   266: 'Carrier 04 Safe Output Card Fault', class No Acknowledgement, trigger "DB302_HMI_Faults_Carrier4_Faults_0" bit 9
   267: 'Carrier 04 Standard Input Card Fault', class No Acknowledgement, trigger "DB302_HMI_Faults_Carrier4_Faults_0" bit 10
   268: 'Carrier 04 Standard Output Card Fault', class No Acknowledgement, trigger "DB302_HMI_Faults_Carrier4_Faults_0" bit 11
   269: 'Carrier 04 Encoder Position Fault', class No Acknowledgement, trigger "DB302_HMI_Faults_Carrier4_Faults_0" bit 12
   270: 'Carrier 04 Encoder Internal Error', class No Acknowledgement, trigger "DB302_HMI_Faults_Carrier4_Faults_0" bit 13
   271: 'Carrier 04 Encoder Comm Fault', class No Acknowledgement, trigger "DB302_HMI_Faults_Carrier4_Faults_0" bit 14
   272: 'Carrier 04 HMI Comm Fault', class No Acknowledgement, trigger "DB302_HMI_Faults_Carrier4_Faults_0" bit 15
   273: 'Carrier 04 Crash Detection Fault', class No Acknowledgement, trigger "DB302_HMI_Faults_Carrier4_Faults_1" bit 0
   274: 'Carrier 04 Carrier Number Invalid', class No Acknowledgement, trigger "DB302_HMI_Faults_Carrier4_Faults_1" bit 1
   275: 'Carrier 04 Drive: PROFINET configuration error', class No Acknowledgement, trigger "DB302_HMI_Faults_Carrier4_Faults_1" bit 2
   276: 'Carrier 04 Drive: Error internal communications', class No Acknowledgement, trigger "DB302_HMI_Faults_Carrier4_Faults_1" bit 3
   277: 'Carrier 04 Drive: Motor overtemperature', class No Acknowledgement, trigger "DB302_HMI_Faults_Carrier4_Faults_1" bit 4
   278: 'Carrier 04 Drive: Motor overcurrent', class No Acknowledgement, trigger "DB302_HMI_Faults_Carrier4_Faults_1" bit 5
   279: 'Carrier 04 Drive: Infeed or power unit not ready', class No Acknowledgement, trigger "DB302_HMI_Faults_Carrier4_Faults_1" bit 6
   280: 'Carrier 04 Drive: Short-circuit/ground fault detected', class No Acknowledgement, trigger "DB302_HMI_Faults_Carrier4_Faults_1" bit 7
   281: 'Carrier 04 Drive: PROFINET Setpoint timeout', class No Acknowledgement, trigger "DB302_HMI_Faults_Carrier4_Faults_1" bit 8
   282: 'Carrier 04 Power unit: Overcurrent', class No Acknowledgement, trigger "DB302_HMI_Faults_Carrier4_Faults_1" bit 9
   283: 'Carrier 04 Power unit: DC link voltage overvoltage', class No Acknowledgement, trigger "DB302_HMI_Faults_Carrier4_Faults_1" bit 10
   284: 'Carrier 04 Power unit: DC link voltage undervoltage', class No Acknowledgement, trigger "DB302_HMI_Faults_Carrier4_Faults_1" bit 11
   285: 'Carrier 04 Power unit: Line phase failure in main circuit', class No Acknowledgement, trigger "DB302_HMI_Faults_Carrier4_Faults_1" bit 12
   286: 'Carrier 04 Power unit: Phase failure motor cable', class No Acknowledgement, trigger "DB302_HMI_Faults_Carrier4_Faults_1" bit 13
   287: 'Carrier 04 Power unit: Ground fault', class No Acknowledgement, trigger "DB302_HMI_Faults_Carrier4_Faults_1" bit 14
   288: 'Spare_Fault_288', class No Acknowledgement, trigger "DB302_HMI_Faults_Carrier4_Faults_1" bit 15
   289: 'Carrier 04 Motion Off Fault', class No Acknowledgement, trigger "DB302_HMI_Faults_Carrier4_Faults_2" bit 0
   290: 'Carrier 04 Motion On Fault', class No Acknowledgement, trigger "DB302_HMI_Faults_Carrier4_Faults_2" bit 1
   291: 'Carrier 04 Spacing Fault', class No Acknowledgement, trigger "DB302_HMI_Faults_Carrier4_Faults_2" bit 2
   292: 'Carrier 04 Duplicate Carrier Number Fault', class No Acknowledgement, trigger "DB302_HMI_Faults_Carrier4_Faults_2" bit 3
   293: 'Spare_Fault_293', class No Acknowledgement, trigger "DB302_HMI_Faults_Carrier4_Faults_2" bit 4
   294: 'Spare_Fault_294', class No Acknowledgement, trigger "DB302_HMI_Faults_Carrier4_Faults_2" bit 5
   295: 'Spare_Fault_295', class No Acknowledgement, trigger "DB302_HMI_Faults_Carrier4_Faults_2" bit 6
   296: 'Spare_Fault_296', class No Acknowledgement, trigger "DB302_HMI_Faults_Carrier4_Faults_2" bit 7
   297: 'Spare_Fault_297', class No Acknowledgement, trigger "DB302_HMI_Faults_Carrier4_Faults_2" bit 8
   298: 'Spare_Fault_298', class No Acknowledgement, trigger "DB302_HMI_Faults_Carrier4_Faults_2" bit 9
   299: 'Spare_Fault_299', class No Acknowledgement, trigger "DB302_HMI_Faults_Carrier4_Faults_2" bit 10
   300: 'Spare_Fault_300', class No Acknowledgement, trigger "DB302_HMI_Faults_Carrier4_Faults_2" bit 11
   301: 'Spare_Fault_301', class No Acknowledgement, trigger "DB302_HMI_Faults_Carrier4_Faults_2" bit 12
   302: 'Spare_Fault_302', class No Acknowledgement, trigger "DB302_HMI_Faults_Carrier4_Faults_2" bit 13
   303: 'Spare_Fault_303', class No Acknowledgement, trigger "DB302_HMI_Faults_Carrier4_Faults_2" bit 14
   304: 'Spare_Fault_304', class No Acknowledgement, trigger "DB302_HMI_Faults_Carrier4_Faults_2" bit 15
   305: 'Spare_Fault_305', class No Acknowledgement, trigger "DB302_HMI_Faults_Carrier4_Faults_3" bit 0
   306: 'Spare_Fault_306', class No Acknowledgement, trigger "DB302_HMI_Faults_Carrier4_Faults_3" bit 1
   307: 'Spare_Fault_307', class No Acknowledgement, trigger "DB302_HMI_Faults_Carrier4_Faults_3" bit 2
   308: 'Spare_Fault_308', class No Acknowledgement, trigger "DB302_HMI_Faults_Carrier4_Faults_3" bit 3
   309: 'Spare_Fault_309', class No Acknowledgement, trigger "DB302_HMI_Faults_Carrier4_Faults_3" bit 4
   310: 'Spare_Fault_310', class No Acknowledgement, trigger "DB302_HMI_Faults_Carrier4_Faults_3" bit 5
   311: 'Spare_Fault_311', class No Acknowledgement, trigger "DB302_HMI_Faults_Carrier4_Faults_3" bit 6
   312: 'Spare_Fault_312', class No Acknowledgement, trigger "DB302_HMI_Faults_Carrier4_Faults_3" bit 7
   313: 'Spare_Fault_313', class No Acknowledgement, trigger "DB302_HMI_Faults_Carrier4_Faults_3" bit 8
   314: 'Spare_Fault_314', class No Acknowledgement, trigger "DB302_HMI_Faults_Carrier4_Faults_3" bit 9
   315: 'Spare_Fault_315', class No Acknowledgement, trigger "DB302_HMI_Faults_Carrier4_Faults_3" bit 10
   316: 'Spare_Fault_316', class No Acknowledgement, trigger "DB302_HMI_Faults_Carrier4_Faults_3" bit 11
   317: 'Spare_Fault_317', class No Acknowledgement, trigger "DB302_HMI_Faults_Carrier4_Faults_3" bit 12
   318: 'Spare_Fault_318', class No Acknowledgement, trigger "DB302_HMI_Faults_Carrier4_Faults_3" bit 13
   319: 'Spare_Fault_319', class No Acknowledgement, trigger "DB302_HMI_Faults_Carrier4_Faults_3" bit 14
   320: 'Spare_Fault_320', class No Acknowledgement, trigger "DB302_HMI_Faults_Carrier4_Faults_3" bit 15
   321: 'Carrier 05 Disconnect Open Power Fault DI11.0', class No Acknowledgement, trigger "DB302_HMI_Faults_Carrier5_Faults_0" bit 0
   322: 'Carrier 05 Drive Profinet Comm Fault', class No Acknowledgement, trigger "DB302_HMI_Faults_Carrier5_Faults_0" bit 1
   323: 'Carrier 05 Production Stop Not Reset', class No Acknowledgement, trigger "DB302_HMI_Faults_Carrier5_Faults_0" bit 2
   324: 'Carrier 05 CB02122 Tripped', class No Acknowledgement, trigger "DB302_HMI_Faults_Carrier5_Faults_0" bit 3
   325: 'Carrier 05 CB02123 Tripped', class No Acknowledgement, trigger "DB302_HMI_Faults_Carrier5_Faults_0" bit 4
   326: 'Carrier 05 AUX1 CB Tripped', class No Acknowledgement, trigger "DB302_HMI_Faults_Carrier5_Faults_0" bit 5
   327: 'Carrier 05 AUX2 CB Tripped', class No Acknowledgement, trigger "DB302_HMI_Faults_Carrier5_Faults_0" bit 6
   328: 'Carrier 05 PLC Not Communicating', class No Acknowledgement, trigger "DB302_HMI_Faults_Carrier5_Faults_0" bit 7
   329: 'Carrier 05 Safe Input Card Fault', class No Acknowledgement, trigger "DB302_HMI_Faults_Carrier5_Faults_0" bit 8
   330: 'Carrier 05 Safe Output Card Fault', class No Acknowledgement, trigger "DB302_HMI_Faults_Carrier5_Faults_0" bit 9
   331: 'Carrier 05 Standard Input Card Fault', class No Acknowledgement, trigger "DB302_HMI_Faults_Carrier5_Faults_0" bit 10
   332: 'Carrier 05 Standard Output Card Fault', class No Acknowledgement, trigger "DB302_HMI_Faults_Carrier5_Faults_0" bit 11
   333: 'Carrier 05 Encoder Position Fault', class No Acknowledgement, trigger "DB302_HMI_Faults_Carrier5_Faults_0" bit 12
   334: 'Carrier 05 Encoder Internal Error', class No Acknowledgement, trigger "DB302_HMI_Faults_Carrier5_Faults_0" bit 13
   335: 'Carrier 05 Encoder Comm Fault', class No Acknowledgement, trigger "DB302_HMI_Faults_Carrier5_Faults_0" bit 14
   336: 'Carrier 05 HMI Comm Fault', class No Acknowledgement, trigger "DB302_HMI_Faults_Carrier5_Faults_0" bit 15
   337: 'Carrier 05 Crash Detection Fault', class No Acknowledgement, trigger "DB302_HMI_Faults_Carrier5_Faults_1" bit 0
   338: 'Carrier 05 Carrier Number Invalid', class No Acknowledgement, trigger "DB302_HMI_Faults_Carrier5_Faults_1" bit 1
   339: 'Carrier 05 Drive: PROFINET configuration error', class No Acknowledgement, trigger "DB302_HMI_Faults_Carrier5_Faults_1" bit 2
   340: 'Carrier 05 Drive: Error internal communications', class No Acknowledgement, trigger "DB302_HMI_Faults_Carrier5_Faults_1" bit 3
   341: 'Carrier 05 Drive: Motor overtemperature', class No Acknowledgement, trigger "DB302_HMI_Faults_Carrier5_Faults_1" bit 4
   342: 'Carrier 05 Drive: Motor overcurrent', class No Acknowledgement, trigger "DB302_HMI_Faults_Carrier5_Faults_1" bit 5
   343: 'Carrier 05 Drive: Infeed or power unit not ready', class No Acknowledgement, trigger "DB302_HMI_Faults_Carrier5_Faults_1" bit 6
   344: 'Carrier 05 Drive: Short-circuit/ground fault detected', class No Acknowledgement, trigger "DB302_HMI_Faults_Carrier5_Faults_1" bit 7
   345: 'Carrier 05 Drive: PROFINET Setpoint timeout', class No Acknowledgement, trigger "DB302_HMI_Faults_Carrier5_Faults_1" bit 8
   346: 'Carrier 05 Power unit: Overcurrent', class No Acknowledgement, trigger "DB302_HMI_Faults_Carrier5_Faults_1" bit 9
   347: 'Carrier 05 Power unit: DC link voltage overvoltage', class No Acknowledgement, trigger "DB302_HMI_Faults_Carrier5_Faults_1" bit 10
   348: 'Carrier 05 Power unit: DC link voltage undervoltage', class No Acknowledgement, trigger "DB302_HMI_Faults_Carrier5_Faults_1" bit 11
   349: 'Carrier 05 Power unit: Line phase failure in main circuit', class No Acknowledgement, trigger "DB302_HMI_Faults_Carrier5_Faults_1" bit 12
   350: 'Carrier 05 Power unit: Phase failure motor cable', class No Acknowledgement, trigger "DB302_HMI_Faults_Carrier5_Faults_1" bit 13
   351: 'Carrier 05 Power unit: Ground fault', class No Acknowledgement, trigger "DB302_HMI_Faults_Carrier5_Faults_1" bit 14
   352: 'Spare_Fault_352', class No Acknowledgement, trigger "DB302_HMI_Faults_Carrier5_Faults_1" bit 15
   353: 'Carrier 05 Motion Off Fault', class No Acknowledgement, trigger "DB302_HMI_Faults_Carrier5_Faults_2" bit 0
   354: 'Carrier 05 Motion On Fault', class No Acknowledgement, trigger "DB302_HMI_Faults_Carrier5_Faults_2" bit 1
   355: 'Carrier 05 Spacing Fault', class No Acknowledgement, trigger "DB302_HMI_Faults_Carrier5_Faults_2" bit 2
   356: 'Carrier 05 Duplicate Carrier Number Fault', class No Acknowledgement, trigger "DB302_HMI_Faults_Carrier5_Faults_2" bit 3
   357: 'Spare_Fault_357', class No Acknowledgement, trigger "DB302_HMI_Faults_Carrier5_Faults_2" bit 4
   358: 'Spare_Fault_358', class No Acknowledgement, trigger "DB302_HMI_Faults_Carrier5_Faults_2" bit 5
   359: 'Spare_Fault_359', class No Acknowledgement, trigger "DB302_HMI_Faults_Carrier5_Faults_2" bit 6
   360: 'Spare_Fault_360', class No Acknowledgement, trigger "DB302_HMI_Faults_Carrier5_Faults_2" bit 7
   361: 'Spare_Fault_361', class No Acknowledgement, trigger "DB302_HMI_Faults_Carrier5_Faults_2" bit 8
   362: 'Spare_Fault_362', class No Acknowledgement, trigger "DB302_HMI_Faults_Carrier5_Faults_2" bit 9
   363: 'Spare_Fault_363', class No Acknowledgement, trigger "DB302_HMI_Faults_Carrier5_Faults_2" bit 10
   364: 'Spare_Fault_364', class No Acknowledgement, trigger "DB302_HMI_Faults_Carrier5_Faults_2" bit 11
   365: 'Spare_Fault_365', class No Acknowledgement, trigger "DB302_HMI_Faults_Carrier5_Faults_2" bit 12
   366: 'Spare_Fault_366', class No Acknowledgement, trigger "DB302_HMI_Faults_Carrier5_Faults_2" bit 13
   367: 'Spare_Fault_367', class No Acknowledgement, trigger "DB302_HMI_Faults_Carrier5_Faults_2" bit 14
   368: 'Spare_Fault_368', class No Acknowledgement, trigger "DB302_HMI_Faults_Carrier5_Faults_2" bit 15
   369: 'Spare_Fault_369', class No Acknowledgement, trigger "DB302_HMI_Faults_Carrier5_Faults_3" bit 0
   370: 'Spare_Fault_370', class No Acknowledgement, trigger "DB302_HMI_Faults_Carrier5_Faults_3" bit 1
   371: 'Spare_Fault_371', class No Acknowledgement, trigger "DB302_HMI_Faults_Carrier5_Faults_3" bit 2
   372: 'Spare_Fault_372', class No Acknowledgement, trigger "DB302_HMI_Faults_Carrier5_Faults_3" bit 3
   373: 'Spare_Fault_373', class No Acknowledgement, trigger "DB302_HMI_Faults_Carrier5_Faults_3" bit 4
   374: 'Spare_Fault_374', class No Acknowledgement, trigger "DB302_HMI_Faults_Carrier5_Faults_3" bit 5
   375: 'Spare_Fault_375', class No Acknowledgement, trigger "DB302_HMI_Faults_Carrier5_Faults_3" bit 6
   376: 'Spare_Fault_376', class No Acknowledgement, trigger "DB302_HMI_Faults_Carrier5_Faults_3" bit 7
   377: 'Spare_Fault_377', class No Acknowledgement, trigger "DB302_HMI_Faults_Carrier5_Faults_3" bit 8
   378: 'Spare_Fault_378', class No Acknowledgement, trigger "DB302_HMI_Faults_Carrier5_Faults_3" bit 9
   379: 'Spare_Fault_379', class No Acknowledgement, trigger "DB302_HMI_Faults_Carrier5_Faults_3" bit 10
   380: 'Spare_Fault_380', class No Acknowledgement, trigger "DB302_HMI_Faults_Carrier5_Faults_3" bit 11
   381: 'Spare_Fault_381', class No Acknowledgement, trigger "DB302_HMI_Faults_Carrier5_Faults_3" bit 12
   382: 'Spare_Fault_382', class No Acknowledgement, trigger "DB302_HMI_Faults_Carrier5_Faults_3" bit 13
   383: 'Spare_Fault_383', class No Acknowledgement, trigger "DB302_HMI_Faults_Carrier5_Faults_3" bit 14
   384: 'Spare_Fault_384', class No Acknowledgement, trigger "DB302_HMI_Faults_Carrier5_Faults_3" bit 15
   385: 'Carrier 06 Disconnect Open Power Fault DI11.0', class No Acknowledgement, trigger "DB302_HMI_Faults_Carrier6_Faults_0" bit 0
   386: 'Carrier 06 Drive Profinet Comm Fault', class No Acknowledgement, trigger "DB302_HMI_Faults_Carrier6_Faults_0" bit 1
   387: 'Carrier 06 Production Stop Not Reset', class No Acknowledgement, trigger "DB302_HMI_Faults_Carrier6_Faults_0" bit 2
   388: 'Carrier 06 CB02122 Tripped', class No Acknowledgement, trigger "DB302_HMI_Faults_Carrier6_Faults_0" bit 3
   389: 'Carrier 06 CB02123 Tripped', class No Acknowledgement, trigger "DB302_HMI_Faults_Carrier6_Faults_0" bit 4
   390: 'Carrier 06 AUX1 CB Tripped', class No Acknowledgement, trigger "DB302_HMI_Faults_Carrier6_Faults_0" bit 5
   391: 'Carrier 06 AUX2 CB Tripped', class No Acknowledgement, trigger "DB302_HMI_Faults_Carrier6_Faults_0" bit 6
   392: 'Carrier 06 PLC Not Communicating', class No Acknowledgement, trigger "DB302_HMI_Faults_Carrier6_Faults_0" bit 7
   393: 'Carrier 06 Safe Input Card Fault', class No Acknowledgement, trigger "DB302_HMI_Faults_Carrier6_Faults_0" bit 8
   394: 'Carrier 06 Safe Output Card Fault', class No Acknowledgement, trigger "DB302_HMI_Faults_Carrier6_Faults_0" bit 9
   395: 'Carrier 06 Standard Input Card Fault', class No Acknowledgement, trigger "DB302_HMI_Faults_Carrier6_Faults_0" bit 10
   396: 'Carrier 06 Standard Output Card Fault', class No Acknowledgement, trigger "DB302_HMI_Faults_Carrier6_Faults_0" bit 11
   397: 'Carrier 06 Encoder Position Fault', class No Acknowledgement, trigger "DB302_HMI_Faults_Carrier6_Faults_0" bit 12
   398: 'Carrier 06 Encoder Internal Error', class No Acknowledgement, trigger "DB302_HMI_Faults_Carrier6_Faults_0" bit 13
   399: 'Carrier 06 Encoder Comm Fault', class No Acknowledgement, trigger "DB302_HMI_Faults_Carrier6_Faults_0" bit 14
   400: 'Carrier 06 HMI Comm Fault', class No Acknowledgement, trigger "DB302_HMI_Faults_Carrier6_Faults_0" bit 15
   401: 'Carrier 06 Crash Detection Fault', class No Acknowledgement, trigger "DB302_HMI_Faults_Carrier6_Faults_1" bit 0
   402: 'Carrier 06 Carrier Number Invalid', class No Acknowledgement, trigger "DB302_HMI_Faults_Carrier6_Faults_1" bit 1
   403: 'Carrier 06 Drive: PROFINET configuration error', class No Acknowledgement, trigger "DB302_HMI_Faults_Carrier6_Faults_1" bit 2
   404: 'Carrier 06 Drive: Error internal communications', class No Acknowledgement, trigger "DB302_HMI_Faults_Carrier6_Faults_1" bit 3
   405: 'Carrier 06 Drive: Motor overtemperature', class No Acknowledgement, trigger "DB302_HMI_Faults_Carrier6_Faults_1" bit 4
   406: 'Carrier 06 Drive: Motor overcurrent', class No Acknowledgement, trigger "DB302_HMI_Faults_Carrier6_Faults_1" bit 5
   407: 'Carrier 06 Drive: Infeed or power unit not ready', class No Acknowledgement, trigger "DB302_HMI_Faults_Carrier6_Faults_1" bit 6
   408: 'Carrier 06 Drive: Short-circuit/ground fault detected', class No Acknowledgement, trigger "DB302_HMI_Faults_Carrier6_Faults_1" bit 7
   409: 'Carrier 06 Drive: PROFINET Setpoint timeout', class No Acknowledgement, trigger "DB302_HMI_Faults_Carrier6_Faults_1" bit 8
   410: 'Carrier 06 Power unit: Overcurrent', class No Acknowledgement, trigger "DB302_HMI_Faults_Carrier6_Faults_1" bit 9
   411: 'Carrier 06 Power unit: DC link voltage overvoltage', class No Acknowledgement, trigger "DB302_HMI_Faults_Carrier6_Faults_1" bit 10
   412: 'Carrier 06 Power unit: DC link voltage undervoltage', class No Acknowledgement, trigger "DB302_HMI_Faults_Carrier6_Faults_1" bit 11
   413: 'Carrier 06 Power unit: Line phase failure in main circuit', class No Acknowledgement, trigger "DB302_HMI_Faults_Carrier6_Faults_1" bit 12
   414: 'Carrier 06 Power unit: Phase failure motor cable', class No Acknowledgement, trigger "DB302_HMI_Faults_Carrier6_Faults_1" bit 13
   415: 'Carrier 06 Power unit: Ground fault', class No Acknowledgement, trigger "DB302_HMI_Faults_Carrier6_Faults_1" bit 14
   416: 'Spare_Fault_416', class No Acknowledgement, trigger "DB302_HMI_Faults_Carrier6_Faults_1" bit 15
   417: 'Carrier 06 Motion Off Fault', class No Acknowledgement, trigger "DB302_HMI_Faults_Carrier6_Faults_2" bit 0
   418: 'Carrier 06 Motion On Fault', class No Acknowledgement, trigger "DB302_HMI_Faults_Carrier6_Faults_2" bit 1
   419: 'Carrier 06 Spacing Fault', class No Acknowledgement, trigger "DB302_HMI_Faults_Carrier6_Faults_2" bit 2
   420: 'Carrier 06 Duplicate Carrier Number Fault', class No Acknowledgement, trigger "DB302_HMI_Faults_Carrier6_Faults_2" bit 3
   421: 'Spare_Fault_421', class No Acknowledgement, trigger "DB302_HMI_Faults_Carrier6_Faults_2" bit 4
   422: 'Spare_Fault_422', class No Acknowledgement, trigger "DB302_HMI_Faults_Carrier6_Faults_2" bit 5
   423: 'Spare_Fault_423', class No Acknowledgement, trigger "DB302_HMI_Faults_Carrier6_Faults_2" bit 6
   424: 'Spare_Fault_424', class No Acknowledgement, trigger "DB302_HMI_Faults_Carrier6_Faults_2" bit 7
   425: 'Spare_Fault_425', class No Acknowledgement, trigger "DB302_HMI_Faults_Carrier6_Faults_2" bit 8
   426: 'Spare_Fault_426', class No Acknowledgement, trigger "DB302_HMI_Faults_Carrier6_Faults_2" bit 9
   427: 'Spare_Fault_427', class No Acknowledgement, trigger "DB302_HMI_Faults_Carrier6_Faults_2" bit 10
   428: 'Spare_Fault_428', class No Acknowledgement, trigger "DB302_HMI_Faults_Carrier6_Faults_2" bit 11
   429: 'Spare_Fault_429', class No Acknowledgement, trigger "DB302_HMI_Faults_Carrier6_Faults_2" bit 12
   430: 'Spare_Fault_430', class No Acknowledgement, trigger "DB302_HMI_Faults_Carrier6_Faults_2" bit 13
   431: 'Spare_Fault_431', class No Acknowledgement, trigger "DB302_HMI_Faults_Carrier6_Faults_2" bit 14
   432: 'Spare_Fault_432', class No Acknowledgement, trigger "DB302_HMI_Faults_Carrier6_Faults_2" bit 15
   433: 'Spare_Fault_433', class No Acknowledgement, trigger "DB302_HMI_Faults_Carrier6_Faults_3" bit 0
   434: 'Spare_Fault_434', class No Acknowledgement, trigger "DB302_HMI_Faults_Carrier6_Faults_3" bit 1
   435: 'Spare_Fault_435', class No Acknowledgement, trigger "DB302_HMI_Faults_Carrier6_Faults_3" bit 2
   436: 'Spare_Fault_436', class No Acknowledgement, trigger "DB302_HMI_Faults_Carrier6_Faults_3" bit 3
   437: 'Spare_Fault_437', class No Acknowledgement, trigger "DB302_HMI_Faults_Carrier6_Faults_3" bit 4
   438: 'Spare_Fault_438', class No Acknowledgement, trigger "DB302_HMI_Faults_Carrier6_Faults_3" bit 5
   439: 'Spare_Fault_439', class No Acknowledgement, trigger "DB302_HMI_Faults_Carrier6_Faults_3" bit 6
   440: 'Spare_Fault_440', class No Acknowledgement, trigger "DB302_HMI_Faults_Carrier6_Faults_3" bit 7
   441: 'Spare_Fault_441', class No Acknowledgement, trigger "DB302_HMI_Faults_Carrier6_Faults_3" bit 8
   442: 'Spare_Fault_442', class No Acknowledgement, trigger "DB302_HMI_Faults_Carrier6_Faults_3" bit 9
   443: 'Spare_Fault_443', class No Acknowledgement, trigger "DB302_HMI_Faults_Carrier6_Faults_3" bit 10
   444: 'Spare_Fault_444', class No Acknowledgement, trigger "DB302_HMI_Faults_Carrier6_Faults_3" bit 11
   445: 'Spare_Fault_445', class No Acknowledgement, trigger "DB302_HMI_Faults_Carrier6_Faults_3" bit 12
   446: 'Spare_Fault_446', class No Acknowledgement, trigger "DB302_HMI_Faults_Carrier6_Faults_3" bit 13
   447: 'Spare_Fault_447', class No Acknowledgement, trigger "DB302_HMI_Faults_Carrier6_Faults_3" bit 14
   448: 'Spare_Fault_448', class No Acknowledgement, trigger "DB302_HMI_Faults_Carrier6_Faults_3" bit 15
   449: 'Carrier 07 Disconnect Open Power Fault DI11.0', class No Acknowledgement, trigger "DB302_HMI_Faults_Carrier7_Faults_0" bit 0
   450: 'Carrier 07 Drive Profinet Comm Fault', class No Acknowledgement, trigger "DB302_HMI_Faults_Carrier7_Faults_0" bit 1
   451: 'Carrier 07 Production Stop Not Reset', class No Acknowledgement, trigger "DB302_HMI_Faults_Carrier7_Faults_0" bit 2
   452: 'Carrier 07 CB02122 Tripped', class No Acknowledgement, trigger "DB302_HMI_Faults_Carrier7_Faults_0" bit 3
   453: 'Carrier 07 CB02123 Tripped', class No Acknowledgement, trigger "DB302_HMI_Faults_Carrier7_Faults_0" bit 4
   454: 'Carrier 07 AUX1 CB Tripped', class No Acknowledgement, trigger "DB302_HMI_Faults_Carrier7_Faults_0" bit 5
   455: 'Carrier 07 AUX2 CB Tripped', class No Acknowledgement, trigger "DB302_HMI_Faults_Carrier7_Faults_0" bit 6
   456: 'Carrier 07 PLC Not Communicating', class No Acknowledgement, trigger "DB302_HMI_Faults_Carrier7_Faults_0" bit 7
   457: 'Carrier 07 Safe Input Card Fault', class No Acknowledgement, trigger "DB302_HMI_Faults_Carrier7_Faults_0" bit 8
   458: 'Carrier 07 Safe Output Card Fault', class No Acknowledgement, trigger "DB302_HMI_Faults_Carrier7_Faults_0" bit 9
   459: 'Carrier 07 Standard Input Card Fault', class No Acknowledgement, trigger "DB302_HMI_Faults_Carrier7_Faults_0" bit 10
   460: 'Carrier 07 Standard Output Card Fault', class No Acknowledgement, trigger "DB302_HMI_Faults_Carrier7_Faults_0" bit 11
   461: 'Carrier 07 Encoder Position Fault', class No Acknowledgement, trigger "DB302_HMI_Faults_Carrier7_Faults_0" bit 12
   462: 'Carrier 07 Encoder Internal Error', class No Acknowledgement, trigger "DB302_HMI_Faults_Carrier7_Faults_0" bit 13
   463: 'Carrier 07 Encoder Comm Fault', class No Acknowledgement, trigger "DB302_HMI_Faults_Carrier7_Faults_0" bit 14
   464: 'Carrier 07 HMI Comm Fault', class No Acknowledgement, trigger "DB302_HMI_Faults_Carrier7_Faults_0" bit 15
   465: 'Carrier 07 Crash Detection Fault', class No Acknowledgement, trigger "DB302_HMI_Faults_Carrier7_Faults_1" bit 0
   466: 'Carrier 07 Carrier Number Invalid', class No Acknowledgement, trigger "DB302_HMI_Faults_Carrier7_Faults_1" bit 1
   467: 'Carrier 07 Drive: PROFINET configuration error', class No Acknowledgement, trigger "DB302_HMI_Faults_Carrier7_Faults_1" bit 2
   468: 'Carrier 07 Drive: Error internal communications', class No Acknowledgement, trigger "DB302_HMI_Faults_Carrier7_Faults_1" bit 3
   469: 'Carrier 07 Drive: Motor overtemperature', class No Acknowledgement, trigger "DB302_HMI_Faults_Carrier7_Faults_1" bit 4
   470: 'Carrier 07 Drive: Motor overcurrent', class No Acknowledgement, trigger "DB302_HMI_Faults_Carrier7_Faults_1" bit 5
   471: 'Carrier 07 Drive: Infeed or power unit not ready', class No Acknowledgement, trigger "DB302_HMI_Faults_Carrier7_Faults_1" bit 6
   472: 'Carrier 07 Drive: Short-circuit/ground fault detected', class No Acknowledgement, trigger "DB302_HMI_Faults_Carrier7_Faults_1" bit 7
   473: 'Carrier 07 Drive: PROFINET Setpoint timeout', class No Acknowledgement, trigger "DB302_HMI_Faults_Carrier7_Faults_1" bit 8
   474: 'Carrier 07 Power unit: Overcurrent', class No Acknowledgement, trigger "DB302_HMI_Faults_Carrier7_Faults_1" bit 9
   475: 'Carrier 07 Power unit: DC link voltage overvoltage', class No Acknowledgement, trigger "DB302_HMI_Faults_Carrier7_Faults_1" bit 10
   476: 'Carrier 07 Power unit: DC link voltage undervoltage', class No Acknowledgement, trigger "DB302_HMI_Faults_Carrier7_Faults_1" bit 11
   477: 'Carrier 07 Power unit: Line phase failure in main circuit', class No Acknowledgement, trigger "DB302_HMI_Faults_Carrier7_Faults_1" bit 12
   478: 'Carrier 07 Power unit: Phase failure motor cable', class No Acknowledgement, trigger "DB302_HMI_Faults_Carrier7_Faults_1" bit 13
   479: 'Carrier 07 Power unit: Ground fault', class No Acknowledgement, trigger "DB302_HMI_Faults_Carrier7_Faults_1" bit 14
   480: 'Spare_Fault_480', class No Acknowledgement, trigger "DB302_HMI_Faults_Carrier7_Faults_1" bit 15
   481: 'Carrier 07 Motion Off Fault', class No Acknowledgement, trigger "DB302_HMI_Faults_Carrier7_Faults_2" bit 0
   482: 'Carrier 07 Motion On Fault', class No Acknowledgement, trigger "DB302_HMI_Faults_Carrier7_Faults_2" bit 1
   483: 'Carrier 07 Spacing Fault', class No Acknowledgement, trigger "DB302_HMI_Faults_Carrier7_Faults_2" bit 2
   484: 'Carrier 07 Duplicate Carrier Number Fault', class No Acknowledgement, trigger "DB302_HMI_Faults_Carrier7_Faults_2" bit 3
   485: 'Spare_Fault_485', class No Acknowledgement, trigger "DB302_HMI_Faults_Carrier7_Faults_2" bit 4
   486: 'Spare_Fault_486', class No Acknowledgement, trigger "DB302_HMI_Faults_Carrier7_Faults_2" bit 5
   487: 'Spare_Fault_487', class No Acknowledgement, trigger "DB302_HMI_Faults_Carrier7_Faults_2" bit 6
   488: 'Spare_Fault_488', class No Acknowledgement, trigger "DB302_HMI_Faults_Carrier7_Faults_2" bit 7
   489: 'Spare_Fault_489', class No Acknowledgement, trigger "DB302_HMI_Faults_Carrier7_Faults_2" bit 8
   490: 'Spare_Fault_490', class No Acknowledgement, trigger "DB302_HMI_Faults_Carrier7_Faults_2" bit 9
   491: 'Spare_Fault_491', class No Acknowledgement, trigger "DB302_HMI_Faults_Carrier7_Faults_2" bit 10
   492: 'Spare_Fault_492', class No Acknowledgement, trigger "DB302_HMI_Faults_Carrier7_Faults_2" bit 11
   493: 'Spare_Fault_493', class No Acknowledgement, trigger "DB302_HMI_Faults_Carrier7_Faults_2" bit 12
   494: 'Spare_Fault_494', class No Acknowledgement, trigger "DB302_HMI_Faults_Carrier7_Faults_2" bit 13
   495: 'Spare_Fault_495', class No Acknowledgement, trigger "DB302_HMI_Faults_Carrier7_Faults_2" bit 14
   496: 'Spare_Fault_496', class No Acknowledgement, trigger "DB302_HMI_Faults_Carrier7_Faults_2" bit 15
   497: 'Spare_Fault_497', class No Acknowledgement, trigger "DB302_HMI_Faults_Carrier7_Faults_3" bit 0
   498: 'Spare_Fault_498', class No Acknowledgement, trigger "DB302_HMI_Faults_Carrier7_Faults_3" bit 1
   499: 'Spare_Fault_499', class No Acknowledgement, trigger "DB302_HMI_Faults_Carrier7_Faults_3" bit 2
   500: 'Spare_Fault_500', class No Acknowledgement, trigger "DB302_HMI_Faults_Carrier7_Faults_3" bit 3
   501: 'Spare_Fault_501', class No Acknowledgement, trigger "DB302_HMI_Faults_Carrier7_Faults_3" bit 4
   502: 'Spare_Fault_502', class No Acknowledgement, trigger "DB302_HMI_Faults_Carrier7_Faults_3" bit 5
   503: 'Spare_Fault_503', class No Acknowledgement, trigger "DB302_HMI_Faults_Carrier7_Faults_3" bit 6
   504: 'Spare_Fault_504', class No Acknowledgement, trigger "DB302_HMI_Faults_Carrier7_Faults_3" bit 7
   505: 'Spare_Fault_505', class No Acknowledgement, trigger "DB302_HMI_Faults_Carrier7_Faults_3" bit 8
   506: 'Spare_Fault_506', class No Acknowledgement, trigger "DB302_HMI_Faults_Carrier7_Faults_3" bit 9
   507: 'Spare_Fault_507', class No Acknowledgement, trigger "DB302_HMI_Faults_Carrier7_Faults_3" bit 10
   508: 'Spare_Fault_508', class No Acknowledgement, trigger "DB302_HMI_Faults_Carrier7_Faults_3" bit 11
   509: 'Spare_Fault_509', class No Acknowledgement, trigger "DB302_HMI_Faults_Carrier7_Faults_3" bit 12
   510: 'Spare_Fault_510', class No Acknowledgement, trigger "DB302_HMI_Faults_Carrier7_Faults_3" bit 13
   511: 'Spare_Fault_511', class No Acknowledgement, trigger "DB302_HMI_Faults_Carrier7_Faults_3" bit 14
   512: 'Spare_Fault_512', class No Acknowledgement, trigger "DB302_HMI_Faults_Carrier7_Faults_3" bit 15
   513: 'Carrier 08 Disconnect Open Power Fault DI11.0', class No Acknowledgement, trigger "DB302_HMI_Faults_Carrier8_Faults_0" bit 0
   514: 'Carrier 08 Drive Profinet Comm Fault', class No Acknowledgement, trigger "DB302_HMI_Faults_Carrier8_Faults_0" bit 1
   515: 'Carrier 08 Production Stop Not Reset', class No Acknowledgement, trigger "DB302_HMI_Faults_Carrier8_Faults_0" bit 2
   516: 'Carrier 08 CB02122 Tripped', class No Acknowledgement, trigger "DB302_HMI_Faults_Carrier8_Faults_0" bit 3
   517: 'Carrier 08 CB02123 Tripped', class No Acknowledgement, trigger "DB302_HMI_Faults_Carrier8_Faults_0" bit 4
   518: 'Carrier 08 AUX1 CB Tripped', class No Acknowledgement, trigger "DB302_HMI_Faults_Carrier8_Faults_0" bit 5
   519: 'Carrier 08 AUX2 CB Tripped', class No Acknowledgement, trigger "DB302_HMI_Faults_Carrier8_Faults_0" bit 6
   520: 'Carrier 08 PLC Not Communicating', class No Acknowledgement, trigger "DB302_HMI_Faults_Carrier8_Faults_0" bit 7
   521: 'Carrier 08 Safe Input Card Fault', class No Acknowledgement, trigger "DB302_HMI_Faults_Carrier8_Faults_0" bit 8
   522: 'Carrier 08 Safe Output Card Fault', class No Acknowledgement, trigger "DB302_HMI_Faults_Carrier8_Faults_0" bit 9
   523: 'Carrier 08 Standard Input Card Fault', class No Acknowledgement, trigger "DB302_HMI_Faults_Carrier8_Faults_0" bit 10
   524: 'Carrier 08 Standard Output Card Fault', class No Acknowledgement, trigger "DB302_HMI_Faults_Carrier8_Faults_0" bit 11
   525: 'Carrier 08 Encoder Position Fault', class No Acknowledgement, trigger "DB302_HMI_Faults_Carrier8_Faults_0" bit 12
   526: 'Carrier 08 Encoder Internal Error', class No Acknowledgement, trigger "DB302_HMI_Faults_Carrier8_Faults_0" bit 13
   527: 'Carrier 08 Encoder Comm Fault', class No Acknowledgement, trigger "DB302_HMI_Faults_Carrier8_Faults_0" bit 14
   528: 'Carrier 08 HMI Comm Fault', class No Acknowledgement, trigger "DB302_HMI_Faults_Carrier8_Faults_0" bit 15
   529: 'Carrier 08 Crash Detection Fault', class No Acknowledgement, trigger "DB302_HMI_Faults_Carrier8_Faults_1" bit 0
   530: 'Carrier 08 Carrier Number Invalid', class No Acknowledgement, trigger "DB302_HMI_Faults_Carrier8_Faults_1" bit 1
   531: 'Carrier 08 Drive: PROFINET configuration error', class No Acknowledgement, trigger "DB302_HMI_Faults_Carrier8_Faults_1" bit 2
   532: 'Carrier 08 Drive: Error internal communications', class No Acknowledgement, trigger "DB302_HMI_Faults_Carrier8_Faults_1" bit 3
   533: 'Carrier 08 Drive: Motor overtemperature', class No Acknowledgement, trigger "DB302_HMI_Faults_Carrier8_Faults_1" bit 4
   534: 'Carrier 08 Drive: Motor overcurrent', class No Acknowledgement, trigger "DB302_HMI_Faults_Carrier8_Faults_1" bit 5
   535: 'Carrier 08 Drive: Infeed or power unit not ready', class No Acknowledgement, trigger "DB302_HMI_Faults_Carrier8_Faults_1" bit 6
   536: 'Carrier 08 Drive: Short-circuit/ground fault detected', class No Acknowledgement, trigger "DB302_HMI_Faults_Carrier8_Faults_1" bit 7
   537: 'Carrier 08 Drive: PROFINET Setpoint timeout', class No Acknowledgement, trigger "DB302_HMI_Faults_Carrier8_Faults_1" bit 8
   538: 'Carrier 08 Power unit: Overcurrent', class No Acknowledgement, trigger "DB302_HMI_Faults_Carrier8_Faults_1" bit 9
   539: 'Carrier 08 Power unit: DC link voltage overvoltage', class No Acknowledgement, trigger "DB302_HMI_Faults_Carrier8_Faults_1" bit 10
   540: 'Carrier 08 Power unit: DC link voltage undervoltage', class No Acknowledgement, trigger "DB302_HMI_Faults_Carrier8_Faults_1" bit 11
   541: 'Carrier 08 Power unit: Line phase failure in main circuit', class No Acknowledgement, trigger "DB302_HMI_Faults_Carrier8_Faults_1" bit 12
   542: 'Carrier 08 Power unit: Phase failure motor cable', class No Acknowledgement, trigger "DB302_HMI_Faults_Carrier8_Faults_1" bit 13
   543: 'Carrier 08 Power unit: Ground fault', class No Acknowledgement, trigger "DB302_HMI_Faults_Carrier8_Faults_1" bit 14
   544: 'Spare_Fault_544', class No Acknowledgement, trigger "DB302_HMI_Faults_Carrier8_Faults_1" bit 15
   545: 'Carrier 08 Motion Off Fault', class No Acknowledgement, trigger "DB302_HMI_Faults_Carrier8_Faults_2" bit 0
   546: 'Carrier 08 Motion On Fault', class No Acknowledgement, trigger "DB302_HMI_Faults_Carrier8_Faults_2" bit 1
   547: 'Carrier 08 Spacing Fault', class No Acknowledgement, trigger "DB302_HMI_Faults_Carrier8_Faults_2" bit 2
   548: 'Carrier 08 Duplicate Carrier Number Fault', class No Acknowledgement, trigger "DB302_HMI_Faults_Carrier8_Faults_2" bit 3
   549: 'Spare_Fault_549', class No Acknowledgement, trigger "DB302_HMI_Faults_Carrier8_Faults_2" bit 4
   550: 'Spare_Fault_550', class No Acknowledgement, trigger "DB302_HMI_Faults_Carrier8_Faults_2" bit 5
   551: 'Spare_Fault_551', class No Acknowledgement, trigger "DB302_HMI_Faults_Carrier8_Faults_2" bit 6
   552: 'Spare_Fault_552', class No Acknowledgement, trigger "DB302_HMI_Faults_Carrier8_Faults_2" bit 7
   553: 'Spare_Fault_553', class No Acknowledgement, trigger "DB302_HMI_Faults_Carrier8_Faults_2" bit 8
   554: 'Spare_Fault_554', class No Acknowledgement, trigger "DB302_HMI_Faults_Carrier8_Faults_2" bit 9
   555: 'Spare_Fault_555', class No Acknowledgement, trigger "DB302_HMI_Faults_Carrier8_Faults_2" bit 10
   556: 'Spare_Fault_556', class No Acknowledgement, trigger "DB302_HMI_Faults_Carrier8_Faults_2" bit 11
   557: 'Spare_Fault_557', class No Acknowledgement, trigger "DB302_HMI_Faults_Carrier8_Faults_2" bit 12
   558: 'Spare_Fault_558', class No Acknowledgement, trigger "DB302_HMI_Faults_Carrier8_Faults_2" bit 13
   559: 'Spare_Fault_559', class No Acknowledgement, trigger "DB302_HMI_Faults_Carrier8_Faults_2" bit 14
   560: 'Spare_Fault_560', class No Acknowledgement, trigger "DB302_HMI_Faults_Carrier8_Faults_2" bit 15
   561: 'Spare_Fault_561', class No Acknowledgement, trigger "DB302_HMI_Faults_Carrier8_Faults_3" bit 0
   562: 'Spare_Fault_562', class No Acknowledgement, trigger "DB302_HMI_Faults_Carrier8_Faults_3" bit 1
   563: 'Spare_Fault_563', class No Acknowledgement, trigger "DB302_HMI_Faults_Carrier8_Faults_3" bit 2
   564: 'Spare_Fault_564', class No Acknowledgement, trigger "DB302_HMI_Faults_Carrier8_Faults_3" bit 3
   565: 'Spare_Fault_565', class No Acknowledgement, trigger "DB302_HMI_Faults_Carrier8_Faults_3" bit 4
   566: 'Spare_Fault_566', class No Acknowledgement, trigger "DB302_HMI_Faults_Carrier8_Faults_3" bit 5
   567: 'Spare_Fault_567', class No Acknowledgement, trigger "DB302_HMI_Faults_Carrier8_Faults_3" bit 6
   568: 'Spare_Fault_568', class No Acknowledgement, trigger "DB302_HMI_Faults_Carrier8_Faults_3" bit 7
   569: 'Spare_Fault_569', class No Acknowledgement, trigger "DB302_HMI_Faults_Carrier8_Faults_3" bit 8
   570: 'Spare_Fault_570', class No Acknowledgement, trigger "DB302_HMI_Faults_Carrier8_Faults_3" bit 9
   571: 'Spare_Fault_571', class No Acknowledgement, trigger "DB302_HMI_Faults_Carrier8_Faults_3" bit 10
   572: 'Spare_Fault_572', class No Acknowledgement, trigger "DB302_HMI_Faults_Carrier8_Faults_3" bit 11
   573: 'Spare_Fault_573', class No Acknowledgement, trigger "DB302_HMI_Faults_Carrier8_Faults_3" bit 12
   574: 'Spare_Fault_574', class No Acknowledgement, trigger "DB302_HMI_Faults_Carrier8_Faults_3" bit 13
   575: 'Spare_Fault_575', class No Acknowledgement, trigger "DB302_HMI_Faults_Carrier8_Faults_3" bit 14
   576: 'Spare_Fault_576', class No Acknowledgement, trigger "DB302_HMI_Faults_Carrier8_Faults_3" bit 15
   577: 'Carrier 09 Disconnect Open Power Fault DI11.0', class No Acknowledgement, trigger "DB302_HMI_Faults_Carrier9_Faults_0" bit 0
   578: 'Carrier 09 Drive Profinet Comm Fault', class No Acknowledgement, trigger "DB302_HMI_Faults_Carrier9_Faults_0" bit 1
   579: 'Carrier 09 Production Stop Not Reset', class No Acknowledgement, trigger "DB302_HMI_Faults_Carrier9_Faults_0" bit 2
   580: 'Carrier 09 CB02122 Tripped', class No Acknowledgement, trigger "DB302_HMI_Faults_Carrier9_Faults_0" bit 3
   581: 'Carrier 09 CB02123 Tripped', class No Acknowledgement, trigger "DB302_HMI_Faults_Carrier9_Faults_0" bit 4
   582: 'Carrier 09 AUX1 CB Tripped', class No Acknowledgement, trigger "DB302_HMI_Faults_Carrier9_Faults_0" bit 5
   583: 'Carrier 09 AUX2 CB Tripped', class No Acknowledgement, trigger "DB302_HMI_Faults_Carrier9_Faults_0" bit 6
   584: 'Carrier 09 PLC Not Communicating', class No Acknowledgement, trigger "DB302_HMI_Faults_Carrier9_Faults_0" bit 7
   585: 'Carrier 09 Safe Input Card Fault', class No Acknowledgement, trigger "DB302_HMI_Faults_Carrier9_Faults_0" bit 8
   586: 'Carrier 09 Safe Output Card Fault', class No Acknowledgement, trigger "DB302_HMI_Faults_Carrier9_Faults_0" bit 9
   587: 'Carrier 09 Standard Input Card Fault', class No Acknowledgement, trigger "DB302_HMI_Faults_Carrier9_Faults_0" bit 10
   588: 'Carrier 09 Standard Output Card Fault', class No Acknowledgement, trigger "DB302_HMI_Faults_Carrier9_Faults_0" bit 11
   589: 'Carrier 09 Encoder Position Fault', class No Acknowledgement, trigger "DB302_HMI_Faults_Carrier9_Faults_0" bit 12
   590: 'Carrier 09 Encoder Internal Error', class No Acknowledgement, trigger "DB302_HMI_Faults_Carrier9_Faults_0" bit 13
   591: 'Carrier 09 Encoder Comm Fault', class No Acknowledgement, trigger "DB302_HMI_Faults_Carrier9_Faults_0" bit 14
   592: 'Carrier 09 HMI Comm Fault', class No Acknowledgement, trigger "DB302_HMI_Faults_Carrier9_Faults_0" bit 15
   593: 'Carrier 09 Crash Detection Fault', class No Acknowledgement, trigger "DB302_HMI_Faults_Carrier9_Faults_1" bit 0
   594: 'Carrier 09 Carrier Number Invalid', class No Acknowledgement, trigger "DB302_HMI_Faults_Carrier9_Faults_1" bit 1
   595: 'Carrier 09 Drive: PROFINET configuration error', class No Acknowledgement, trigger "DB302_HMI_Faults_Carrier9_Faults_1" bit 2
   596: 'Carrier 09 Drive: Error internal communications', class No Acknowledgement, trigger "DB302_HMI_Faults_Carrier9_Faults_1" bit 3
   597: 'Carrier 09 Drive: Motor overtemperature', class No Acknowledgement, trigger "DB302_HMI_Faults_Carrier9_Faults_1" bit 4
   598: 'Carrier 09 Drive: Motor overcurrent', class No Acknowledgement, trigger "DB302_HMI_Faults_Carrier9_Faults_1" bit 5
   599: 'Carrier 09 Drive: Infeed or power unit not ready', class No Acknowledgement, trigger "DB302_HMI_Faults_Carrier9_Faults_1" bit 6
   600: 'Carrier 09 Drive: Short-circuit/ground fault detected', class No Acknowledgement, trigger "DB302_HMI_Faults_Carrier9_Faults_1" bit 7
   601: 'Carrier 09 Drive: PROFINET Setpoint timeout', class No Acknowledgement, trigger "DB302_HMI_Faults_Carrier9_Faults_1" bit 8
   602: 'Carrier 09 Power unit: Overcurrent', class No Acknowledgement, trigger "DB302_HMI_Faults_Carrier9_Faults_1" bit 9
   603: 'Carrier 09 Power unit: DC link voltage overvoltage', class No Acknowledgement, trigger "DB302_HMI_Faults_Carrier9_Faults_1" bit 10
   604: 'Carrier 09 Power unit: DC link voltage undervoltage', class No Acknowledgement, trigger "DB302_HMI_Faults_Carrier9_Faults_1" bit 11
   605: 'Carrier 09 Power unit: Line phase failure in main circuit', class No Acknowledgement, trigger "DB302_HMI_Faults_Carrier9_Faults_1" bit 12
   606: 'Carrier 09 Power unit: Phase failure motor cable', class No Acknowledgement, trigger "DB302_HMI_Faults_Carrier9_Faults_1" bit 13
   607: 'Carrier 09 Power unit: Ground fault', class No Acknowledgement, trigger "DB302_HMI_Faults_Carrier9_Faults_1" bit 14
   608: 'Spare_Fault_608', class No Acknowledgement, trigger "DB302_HMI_Faults_Carrier9_Faults_1" bit 15
   609: 'Carrier 09 Motion Off Fault', class No Acknowledgement, trigger "DB302_HMI_Faults_Carrier9_Faults_2" bit 0
   610: 'Carrier 09 Motion On Fault', class No Acknowledgement, trigger "DB302_HMI_Faults_Carrier9_Faults_2" bit 1
   611: 'Carrier 09 Spacing Fault', class No Acknowledgement, trigger "DB302_HMI_Faults_Carrier9_Faults_2" bit 2
   612: 'Carrier 09 Duplicate Carrier Number Fault', class No Acknowledgement, trigger "DB302_HMI_Faults_Carrier9_Faults_2" bit 3
   613: 'Spare_Fault_613', class No Acknowledgement, trigger "DB302_HMI_Faults_Carrier9_Faults_2" bit 4
   614: 'Spare_Fault_614', class No Acknowledgement, trigger "DB302_HMI_Faults_Carrier9_Faults_2" bit 5
   615: 'Spare_Fault_615', class No Acknowledgement, trigger "DB302_HMI_Faults_Carrier9_Faults_2" bit 6
   616: 'Spare_Fault_616', class No Acknowledgement, trigger "DB302_HMI_Faults_Carrier9_Faults_2" bit 7
   617: 'Spare_Fault_617', class No Acknowledgement, trigger "DB302_HMI_Faults_Carrier9_Faults_2" bit 8
   618: 'Spare_Fault_618', class No Acknowledgement, trigger "DB302_HMI_Faults_Carrier9_Faults_2" bit 9
   619: 'Spare_Fault_619', class No Acknowledgement, trigger "DB302_HMI_Faults_Carrier9_Faults_2" bit 10
   620: 'Spare_Fault_620', class No Acknowledgement, trigger "DB302_HMI_Faults_Carrier9_Faults_2" bit 11
   621: 'Spare_Fault_621', class No Acknowledgement, trigger "DB302_HMI_Faults_Carrier9_Faults_2" bit 12
   622: 'Spare_Fault_622', class No Acknowledgement, trigger "DB302_HMI_Faults_Carrier9_Faults_2" bit 13
   623: 'Spare_Fault_623', class No Acknowledgement, trigger "DB302_HMI_Faults_Carrier9_Faults_2" bit 14
   624: 'Spare_Fault_624', class No Acknowledgement, trigger "DB302_HMI_Faults_Carrier9_Faults_2" bit 15
   625: 'Spare_Fault_625', class No Acknowledgement, trigger "DB302_HMI_Faults_Carrier9_Faults_3" bit 0
   626: 'Spare_Fault_626', class No Acknowledgement, trigger "DB302_HMI_Faults_Carrier9_Faults_3" bit 1
   627: 'Spare_Fault_627', class No Acknowledgement, trigger "DB302_HMI_Faults_Carrier9_Faults_3" bit 2
   628: 'Spare_Fault_628', class No Acknowledgement, trigger "DB302_HMI_Faults_Carrier9_Faults_3" bit 3
   629: 'Spare_Fault_629', class No Acknowledgement, trigger "DB302_HMI_Faults_Carrier9_Faults_3" bit 4
   630: 'Spare_Fault_630', class No Acknowledgement, trigger "DB302_HMI_Faults_Carrier9_Faults_3" bit 5
   631: 'Spare_Fault_631', class No Acknowledgement, trigger "DB302_HMI_Faults_Carrier9_Faults_3" bit 6
   632: 'Spare_Fault_632', class No Acknowledgement, trigger "DB302_HMI_Faults_Carrier9_Faults_3" bit 7
   633: 'Spare_Fault_633', class No Acknowledgement, trigger "DB302_HMI_Faults_Carrier9_Faults_3" bit 8
   634: 'Spare_Fault_634', class No Acknowledgement, trigger "DB302_HMI_Faults_Carrier9_Faults_3" bit 9
   635: 'Spare_Fault_635', class No Acknowledgement, trigger "DB302_HMI_Faults_Carrier9_Faults_3" bit 10
   636: 'Spare_Fault_636', class No Acknowledgement, trigger "DB302_HMI_Faults_Carrier9_Faults_3" bit 11
   637: 'Spare_Fault_637', class No Acknowledgement, trigger "DB302_HMI_Faults_Carrier9_Faults_3" bit 12
   638: 'Spare_Fault_638', class No Acknowledgement, trigger "DB302_HMI_Faults_Carrier9_Faults_3" bit 13
   639: 'Spare_Fault_639', class No Acknowledgement, trigger "DB302_HMI_Faults_Carrier9_Faults_3" bit 14
   640: 'Spare_Fault_640', class No Acknowledgement, trigger "DB302_HMI_Faults_Carrier9_Faults_3" bit 15
   641: 'Carrier 10 Disconnect Open Power Fault DI11.0', class No Acknowledgement, trigger "DB302_HMI_Faults_Carrier10_Faults_0" bit 0
   642: 'Carrier 10 Drive Profinet Comm Fault', class No Acknowledgement, trigger "DB302_HMI_Faults_Carrier10_Faults_0" bit 1
   643: 'Carrier 10 Production Stop Not Reset', class No Acknowledgement, trigger "DB302_HMI_Faults_Carrier10_Faults_0" bit 2
   644: 'Carrier 10 CB02122 Tripped', class No Acknowledgement, trigger "DB302_HMI_Faults_Carrier10_Faults_0" bit 3
   645: 'Carrier 10 CB02123 Tripped', class No Acknowledgement, trigger "DB302_HMI_Faults_Carrier10_Faults_0" bit 4
   646: 'Carrier 10 AUX1 CB Tripped', class No Acknowledgement, trigger "DB302_HMI_Faults_Carrier10_Faults_0" bit 5
   647: 'Carrier 10 AUX2 CB Tripped', class No Acknowledgement, trigger "DB302_HMI_Faults_Carrier10_Faults_0" bit 6
   648: 'Carrier 10 PLC Not Communicating', class No Acknowledgement, trigger "DB302_HMI_Faults_Carrier10_Faults_0" bit 7
   649: 'Carrier 10 Safe Input Card Fault', class No Acknowledgement, trigger "DB302_HMI_Faults_Carrier10_Faults_0" bit 8
   650: 'Carrier 10 Safe Output Card Fault', class No Acknowledgement, trigger "DB302_HMI_Faults_Carrier10_Faults_0" bit 9
   651: 'Carrier 10 Standard Input Card Fault', class No Acknowledgement, trigger "DB302_HMI_Faults_Carrier10_Faults_0" bit 10
   652: 'Carrier 10 Standard Output Card Fault', class No Acknowledgement, trigger "DB302_HMI_Faults_Carrier10_Faults_0" bit 11
   653: 'Carrier 10 Encoder Position Fault', class No Acknowledgement, trigger "DB302_HMI_Faults_Carrier10_Faults_0" bit 12
   654: 'Carrier 10 Encoder Internal Error', class No Acknowledgement, trigger "DB302_HMI_Faults_Carrier10_Faults_0" bit 13
   655: 'Carrier 10 Encoder Comm Fault', class No Acknowledgement, trigger "DB302_HMI_Faults_Carrier10_Faults_0" bit 14
   656: 'Carrier 10 HMI Comm Fault', class No Acknowledgement, trigger "DB302_HMI_Faults_Carrier10_Faults_0" bit 15
   657: 'Carrier 10 Crash Detection Fault', class No Acknowledgement, trigger "DB302_HMI_Faults_Carrier10_Faults_1" bit 0
   658: 'Carrier 10 Carrier Number Invalid', class No Acknowledgement, trigger "DB302_HMI_Faults_Carrier10_Faults_1" bit 1
   659: 'Carrier 10 Drive: PROFINET configuration error', class No Acknowledgement, trigger "DB302_HMI_Faults_Carrier10_Faults_1" bit 2
   660: 'Carrier 10 Drive: Error internal communications', class No Acknowledgement, trigger "DB302_HMI_Faults_Carrier10_Faults_1" bit 3
   661: 'Carrier 10 Drive: Motor overtemperature', class No Acknowledgement, trigger "DB302_HMI_Faults_Carrier10_Faults_1" bit 4
   662: 'Carrier 10 Drive: Motor overcurrent', class No Acknowledgement, trigger "DB302_HMI_Faults_Carrier10_Faults_1" bit 5
   663: 'Carrier 10 Drive: Infeed or power unit not ready', class No Acknowledgement, trigger "DB302_HMI_Faults_Carrier10_Faults_1" bit 6
   664: 'Carrier 10 Drive: Short-circuit/ground fault detected', class No Acknowledgement, trigger "DB302_HMI_Faults_Carrier10_Faults_1" bit 7
   665: 'Carrier 10 Drive: PROFINET Setpoint timeout', class No Acknowledgement, trigger "DB302_HMI_Faults_Carrier10_Faults_1" bit 8
   666: 'Carrier 10 Power unit: Overcurrent', class No Acknowledgement, trigger "DB302_HMI_Faults_Carrier10_Faults_1" bit 9
   667: 'Carrier 10 Power unit: DC link voltage overvoltage', class No Acknowledgement, trigger "DB302_HMI_Faults_Carrier10_Faults_1" bit 10
   668: 'Carrier 10 Power unit: DC link voltage undervoltage', class No Acknowledgement, trigger "DB302_HMI_Faults_Carrier10_Faults_1" bit 11
   669: 'Carrier 10 Power unit: Line phase failure in main circuit', class No Acknowledgement, trigger "DB302_HMI_Faults_Carrier10_Faults_1" bit 12
   670: 'Carrier 10 Power unit: Phase failure motor cable', class No Acknowledgement, trigger "DB302_HMI_Faults_Carrier10_Faults_1" bit 13
   671: 'Carrier 10 Power unit: Ground fault', class No Acknowledgement, trigger "DB302_HMI_Faults_Carrier10_Faults_1" bit 14
   672: 'Spare_Fault_672', class No Acknowledgement, trigger "DB302_HMI_Faults_Carrier10_Faults_1" bit 15
   673: 'Carrier 10 Motion Off Fault', class No Acknowledgement, trigger "DB302_HMI_Faults_Carrier10_Faults_2" bit 0
   674: 'Carrier 10 Motion On Fault', class No Acknowledgement, trigger "DB302_HMI_Faults_Carrier10_Faults_2" bit 1
   675: 'Carrier 10 Spacing Fault', class No Acknowledgement, trigger "DB302_HMI_Faults_Carrier10_Faults_2" bit 2
   676: 'Carrier 10 Duplicate Carrier Number Fault', class No Acknowledgement, trigger "DB302_HMI_Faults_Carrier10_Faults_2" bit 3
   677: 'Spare_Fault_677', class No Acknowledgement, trigger "DB302_HMI_Faults_Carrier10_Faults_2" bit 4
   678: 'Spare_Fault_678', class No Acknowledgement, trigger "DB302_HMI_Faults_Carrier10_Faults_2" bit 5
   679: 'Spare_Fault_679', class No Acknowledgement, trigger "DB302_HMI_Faults_Carrier10_Faults_2" bit 6
   680: 'Spare_Fault_680', class No Acknowledgement, trigger "DB302_HMI_Faults_Carrier10_Faults_2" bit 7
   681: 'Spare_Fault_681', class No Acknowledgement, trigger "DB302_HMI_Faults_Carrier10_Faults_2" bit 8
   682: 'Spare_Fault_682', class No Acknowledgement, trigger "DB302_HMI_Faults_Carrier10_Faults_2" bit 9
   683: 'Spare_Fault_683', class No Acknowledgement, trigger "DB302_HMI_Faults_Carrier10_Faults_2" bit 10
   684: 'Spare_Fault_684', class No Acknowledgement, trigger "DB302_HMI_Faults_Carrier10_Faults_2" bit 11
   685: 'Spare_Fault_685', class No Acknowledgement, trigger "DB302_HMI_Faults_Carrier10_Faults_2" bit 12
   686: 'Spare_Fault_686', class No Acknowledgement, trigger "DB302_HMI_Faults_Carrier10_Faults_2" bit 13
   687: 'Spare_Fault_687', class No Acknowledgement, trigger "DB302_HMI_Faults_Carrier10_Faults_2" bit 14
   688: 'Spare_Fault_688', class No Acknowledgement, trigger "DB302_HMI_Faults_Carrier10_Faults_2" bit 15
   689: 'Spare_Fault_689', class No Acknowledgement, trigger "DB302_HMI_Faults_Carrier10_Faults_3" bit 0
   690: 'Spare_Fault_690', class No Acknowledgement, trigger "DB302_HMI_Faults_Carrier10_Faults_3" bit 1
   691: 'Spare_Fault_691', class No Acknowledgement, trigger "DB302_HMI_Faults_Carrier10_Faults_3" bit 2
   692: 'Spare_Fault_692', class No Acknowledgement, trigger "DB302_HMI_Faults_Carrier10_Faults_3" bit 3
   693: 'Spare_Fault_693', class No Acknowledgement, trigger "DB302_HMI_Faults_Carrier10_Faults_3" bit 4
